// TIA Portal project "SWNC V2.0" (V16)

(* hardware
DEVICE "S7-1200 station_1"  S7-1200 Station
   slot 0: "Rack_0"  S7-1200 Rack  Rack  V1.0
   slot 1: "Rupert"  CPU 1214C DC/DC/DC  6ES7 214-1AG40-0XB0  V4.4
   slot 2: "DI 8x24VDC_1"  6ES7 221-1BF32-0XB0  V2.0
   slot 3: "CB 1241 (RS485)"  CB 1241 (RS485)  6ES7 241-1CH30-1XB0  V1.0
   slot 3: "DQ 8xRelay_1"  SM 1222 DQ8 x relay  6ES7 222-1HF32-0XB0  V2.0
   slot 4: "AI 8x13BIT_1"  6ES7 231-4HF32-0XB0  V2.1
   slot 5: "AQ 2x14BIT_1"  SM 1232 AQ2  6ES7 232-4HB32-0XB0  V2.1
DEVICE "HMI_1"  KTP700 Basic PN
   slot 0: "HMI_1"  KTP700 Basic PN  6AV2 123-2GB03-0AX0  16.0.0.0
   slot 1: "HMI_RT_1"  KTP700 Basic PN  6AV2 123-2GB03-0AX0  16.0.0.0
   slot 5: "HMI_1.IE_CP_1"  PROFINET Interface  16.0.0.0
      slot 1: "PROFINET Interface_1"  PROFINET Interface
         slot 1: "Port_1"  Port
*)

// ===== PLC "Rupert"  CPU 1214C DC/DC/DC =====

VAR_GLOBAL   // PLC tag table "Default tag table"
   "System_Byte" AT %MB1000 : Byte;
   "FirstScan" AT %M1000.0 : Bool;
   "DiagStatusUpdate" AT %M1000.1 : Bool;
   "AlwaysTRUE" AT %M1000.2 : Bool;
   "AlwaysFALSE" AT %M1000.3 : Bool;
   "Clock_Byte" AT %MB1001 : Byte;
   "Clock_10Hz" AT %M1001.0 : Bool;
   "Clock_5Hz" AT %M1001.1 : Bool;
   "Clock_2.5Hz" AT %M1001.2 : Bool;
   "Clock_2Hz" AT %M1001.3 : Bool;
   "Clock_1.25Hz" AT %M1001.4 : Bool;
   "Clock_1Hz" AT %M1001.5 : Bool;
   "Clock_0.625Hz" AT %M1001.6 : Bool;
   "Clock_0.5Hz" AT %M1001.7 : Bool;
   "local time conv" AT %MD0 : Time_Of_Day;
   "DN OS1" AT %M4.0 : Bool;
   "temp 3" AT %M4.2 : Bool;
   "DN transition" AT %M4.3 : Bool;
   "PH HOA manual" AT %M4.4 : Bool;   // placeholder for HOA
   "PH HOA Auto" AT %M4.5 : Bool;   // placeholder
END_VAR

VAR_GLOBAL   // PLC tag table "Times"
   "day / night" AT %M0.0 : Bool;   // 1 day, 0 night
   "ND transition" AT %M4.1 : Bool;
END_VAR

VAR_GLOBAL   // PLC tag table "HOA Modes"
   "HOA mode off" AT %M4.6 : Bool;
   "HOA mode manual" AT %M4.7 : Bool;
   "HOA Mode Auto" AT %M5.0 : Bool;
END_VAR

DATA_BLOCK "What time is it_DB"   // DB1
{ S7_Optimized_Access := 'TRUE' }
VERSION : 0.1
// stored: InstanceOfName What time is it
"What time is it"
BEGIN
END_DATA_BLOCK

DATA_BLOCK "HOA_DB"   // DB6
{ S7_Optimized_Access := 'TRUE' }
VERSION : 0.1
// stored: InstanceOfName HOA
"HOA"
BEGIN
END_DATA_BLOCK

DATA_BLOCK "OFF_DB"   // DB7
{ S7_Optimized_Access := 'TRUE' }
VERSION : 0.1
// stored: InstanceOfName OFF
"OFF"
BEGIN
END_DATA_BLOCK

DATA_BLOCK "MANUAL_DB"   // DB8
{ S7_Optimized_Access := 'TRUE' }
VERSION : 0.1
// stored: InstanceOfName MANUAL
"MANUAL"
BEGIN
END_DATA_BLOCK

DATA_BLOCK "AUTO_DB"   // DB9
{ S7_Optimized_Access := 'TRUE' }
VERSION : 0.1
// stored: InstanceOfName AUTO
"AUTO"
BEGIN
END_DATA_BLOCK

// folder: Time

DATA_BLOCK "times list"   // DB2
{ S7_Optimized_Access := 'TRUE' }
VERSION : 0.1
   VAR
      "local time conv" : Time_Of_Day;
      "nightime start" : Time_Of_Day := TOD#16:10:00;
      "nightime end" : Time_Of_Day := TOD#06:00:00;
   END_VAR
BEGIN
END_DATA_BLOCK

// folder: (top level)

FUNCTION_BLOCK "HOA"   // FB2, LAD
{ S7_Optimized_Access := 'TRUE' }
VERSION : 0.1
BEGIN

REGION Network 1
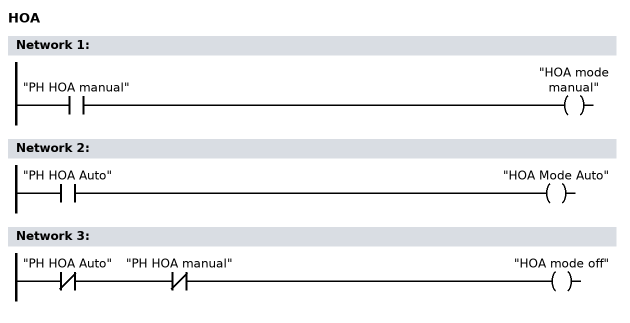
   RUNG wire#powerrail
      Contact( "PH HOA manual" )
      Coil( "HOA mode manual" )
   END_RUNG
   // the same network as SCL:
   "HOA mode manual" := "PH HOA manual";
END_REGION

REGION Network 2
   RUNG wire#powerrail
      Contact( "PH HOA Auto" )
      Coil( "HOA Mode Auto" )
   END_RUNG
   // the same network as SCL:
   "HOA Mode Auto" := "PH HOA Auto";
END_REGION

REGION Network 3
   RUNG wire#powerrail
      I_Contact( "PH HOA Auto" )
      I_Contact( "PH HOA manual" )
      Coil( "HOA mode off" )
   END_RUNG
   // the same network as SCL:
   "HOA mode off" := NOT "PH HOA Auto" AND NOT "PH HOA manual";
END_REGION
END_FUNCTION_BLOCK

ORGANIZATION_BLOCK "Main"   // OB1, LAD, ProgramCycle
TITLE = "Main Program Sweep (Cycle)"
{ S7_Optimized_Access := 'TRUE' }
VERSION : 0.1
   VAR_INPUT
      Initial_Call : Bool;   // Initial call of this OB
      Remanence : Bool;   // =True, if remanent data are available
   END_VAR
BEGIN

REGION Network 1
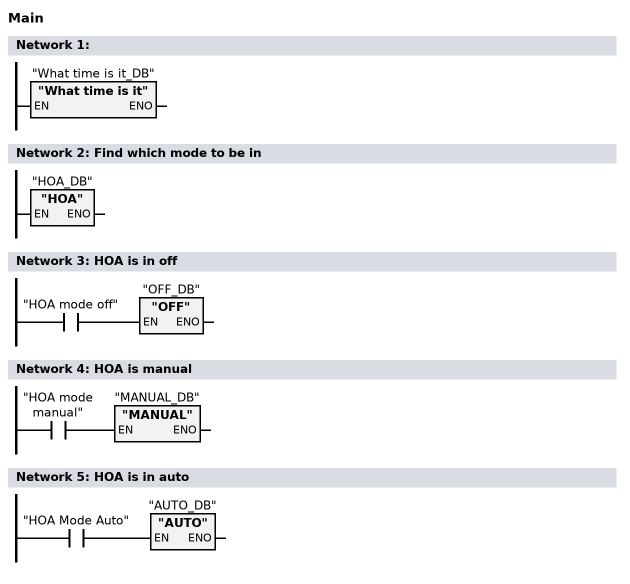
   RUNG wire#powerrail
      "What time is it_DB"()
   END_RUNG
   // the same network as SCL:
   "What time is it_DB"();   // "What time is it"
END_REGION

REGION Network 2: Find which mode to be in
   RUNG wire#powerrail
      "HOA_DB"()
   END_RUNG
   // the same network as SCL:
   "HOA_DB"();   // "HOA"
END_REGION

REGION Network 3: HOA is in off
   RUNG wire#powerrail
      Contact( "HOA mode off" )
      "OFF_DB"()
   END_RUNG
   // the same network as SCL:
   IF "HOA mode off" THEN
       "OFF_DB"();   // "OFF"
   END_IF;
END_REGION

REGION Network 4: HOA is manual
   RUNG wire#powerrail
      Contact( "HOA mode manual" )
      "MANUAL_DB"()
   END_RUNG
   // the same network as SCL:
   IF "HOA mode manual" THEN
       "MANUAL_DB"();   // "MANUAL"
   END_IF;
END_REGION

REGION Network 5: HOA is in auto
   RUNG wire#powerrail
      Contact( "HOA Mode Auto" )
      "AUTO_DB"()
   END_RUNG
   // the same network as SCL:
   IF "HOA Mode Auto" THEN
       "AUTO_DB"();   // "AUTO"
   END_IF;
END_REGION
END_ORGANIZATION_BLOCK

ORGANIZATION_BLOCK "Startup"   // OB100, LAD, Startup
TITLE = "Complete Restart"
{ S7_Optimized_Access := 'TRUE' }
VERSION : 0.1
   VAR_INPUT
      LostRetentive : Bool;   // True if retentive data are lost
      LostRTC : Bool;   // True if date and time are lost
   END_VAR
BEGIN
END_ORGANIZATION_BLOCK

// folder: Modes of operation

FUNCTION_BLOCK "OFF"   // FB3, LAD
{ S7_Optimized_Access := 'TRUE' }
VERSION : 0.1
BEGIN
END_FUNCTION_BLOCK

FUNCTION_BLOCK "AUTO"   // FB4, LAD
{ S7_Optimized_Access := 'TRUE' }
VERSION : 0.1
BEGIN
END_FUNCTION_BLOCK

FUNCTION_BLOCK "MANUAL"   // FB5, LAD
{ S7_Optimized_Access := 'TRUE' }
VERSION : 0.1
BEGIN
END_FUNCTION_BLOCK

// folder: Time

FUNCTION_BLOCK "What time is it"   // FB1, LAD
{ S7_Optimized_Access := 'TRUE' }
VERSION : 0.1
   VAR RETAIN
      "local time" : DTL;
   END_VAR
   VAR
      temp2 : DTL;
      "temp 3" : Bool;
   END_VAR
   VAR_TEMP
      temp : Int;
   END_VAR
   VAR_TEMP   // added for the SCL form of the ladder/FBD networks
      _w1 : Bool;
   END_VAR
BEGIN

REGION Network 1
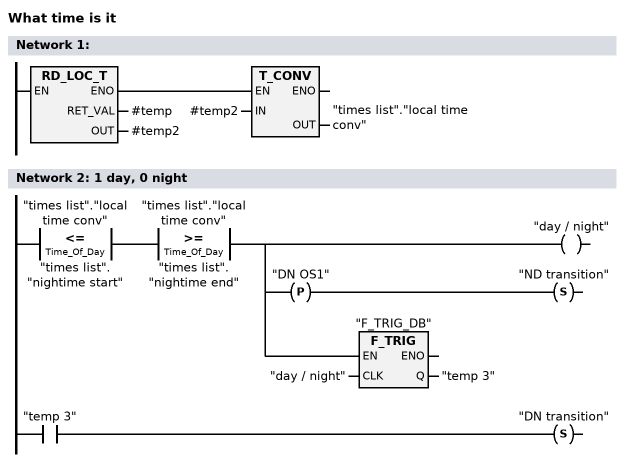
   // ENO of a box is taken as its EN; it also drops when the box reports an error
   #temp := RD_LOC_T(OUT => #temp2);
   "times list"."local time conv" := T_CONV(IN := #temp2);
END_REGION

REGION Network 2: 1 day, 0 night
   "day / night" := ("times list"."local time conv" <= "times list"."nightime start") AND ("times list"."local time conv" >= "times list"."nightime end");
   #_w1 := "day / night" AND NOT "DN OS1";   // rising edge
   "DN OS1" := "day / night";
   IF #_w1 THEN "ND transition" := TRUE; END_IF;
   IF "day / night" THEN
       "F_TRIG_DB"(CLK := "day / night", Q => "temp 3");   // F_TRIG
   END_IF;
   IF "temp 3" THEN "DN transition" := TRUE; END_IF;
END_REGION
END_FUNCTION_BLOCK

(* ===== HMI "HMI_RT_1" =====
system functions are stored by id; their names below are inferred from use
connection "HMI_Connection_1": ETHERNET, SMART_S7_1200_OMS

HMI tags "Default tag table"
   "Tag_ScreenNumber" : UInt, internal

Template "Template_1" 800x480
   Button "Exit" at 714,429 size 71x50; TextOff 'Exit'; PictureOff "ExitRuntime_KTP700_Basic_PN_TR"; PictureOn "ExitRuntime_KTP700_Basic_PN_TR"
      on Release: StopRuntime(0)
   Button "Template_Button" at 614,429 size 71x50; TextOff 'Text'
   Button "Template_Button_1" at 514,429 size 71x50; TextOff 'Text'
   Button "Template_Button_2" at 414,429 size 71x50; TextOff 'Text'
   Button "Template_Button_3" at 314,429 size 71x50; TextOff 'Text'
   Button "Template_Button_4" at 214,429 size 71x50; TextOff 'Text'
   Button "Template_Button_5" at 114,429 size 71x50; TextOff 'Text'
   Button "Start screen" at 14,429 size 71x50; TextOff 'Start screen'; PictureOff "NavigateHome_KTP700_Basic_PN_TR"; PictureOn "NavigateHome_KTP700_Basic_PN_TR"
      on Release: ActivateScreen("Root screen", 0)
   SymbolicIOField "Symbolic_IO_Field_Screen" at 93,9 size 600x33; TextOff '0'; TextOn '1'; TextList "TextList_ScreenNames"
      ProcessValue <- "Tag_ScreenNumber"
      on Change: ActivateScreenByNumber("Tag_ScreenNumber", 0)
   DateTimeField "HmiScreenItemData" at 695,25 size 105x25
   DateTimeField "HmiScreenItemData_1" at 695,0 size 105x25
   GraphicView "Logo" at 0,0 size 91x51; Picture "Logo of HMI_1"

screen "Root screen" 800x480, template "Template_1"
   on GenerateScreen: SetTag("Tag_ScreenNumber", 1)
   TextField "HmiScreenItemData" at 80,225 size 640x25; Text 'Welcome to HMI_1 (KTP700 Basic+ PN)!'
*)